// Mitsubishi GX Works2 project: ZhaoQing_FenRong_Debug   PLC: Q06UDEH (continued)

H750ImportCylinder2(ShuttleCarInOut:= H750ImportCylinder2IO );
ShuttleCarCurrentPosition( XCE OR XCD ,XCE ,XCD, FALSE, H750ImportCylinder2IO.iCurrentPos );
H750ImportCylinder2IO.xReady:=1;
H750ImportCylinder2IO.xForward:=M127;
H750ImportCylinder2IO.xBackward:=M128;
H750ImportCylinder2IO.xPosLimit:=1;
H750ImportCylinder2IO.xNegLimit:=1;
Y2BE:=H750ImportCylinder2IO.xCW;
Y2BD:=H750ImportCylinder2IO.xCCW;
H750ImportCylinder2IO.xCylinder:=1;

H750Conveyor5(ConveyorMotor:=H750Conveyor5IO);
H750Conveyor5IO.xForward:=M112;
H750Conveyor5IO.xCWPresent:=XB6;
Y2AC:=H750Conveyor5IO.xMotorCW;
H750Conveyor5IO.iDeviceID:=12131;

H750Conveyor6(ConveyorMotor:=H750Conveyor6IO);
H750Conveyor6IO.xForward:=M113;
H750Conveyor6IO.xCWPresent:=XB7;
Y2AD:=H750Conveyor6IO.xMotorCW;
H750Conveyor6IO.iDeviceID:=12132;
(********3巷道*************)
H750Switch3(ConveyorEntryIO:=H750Switch3ConveyorIn,
                         ConveyorExitIO:=H750Switch3ConveyorOut,
                        SwitchIO:=H750Switch3IO );
H750Switch3IO.xLiftCylinderExtendButton:=M129;
H750Switch3IO.xLiftCylinderRetractButton:=M130;
H750Switch3IO.xExitBarCylinderRetractButton:=M138;
Y2AF:=NOT (H750Switch3IO.xExitBarCylinderRetract OR m_iH750Switch3Select=2 );
Y2B1:=H750Switch3IO.xLiftCylinderExtend;
Y2B0:=H750Switch3IO.xLiftCylinderRetract;
H750Switch3IO.xLiftCylinderExtendDetect:=XBE;
H750Switch3IO.xLiftCylinderRetractDetect:=XBF;
H750Switch3ConveyorIn.xForward:=M131;
H750Switch3ConveyorIn.xCWPresent:=((m_iH750Switch3Select=1 OR m_iH750Switch3Select=0)  AND  XB9) OR (m_iH750Switch3Select=2 AND XC2);
Y2AB:=H750Switch3ConveyorIn.xMotorCW;
H750Switch3ConveyorIn.tLoadDelay:=T#3s;
H750Switch3ConveyorIn.iDeviceID:=12133;
H750Switch3ConveyorOut.xForward:=M132;
H750Switch3ConveyorOut.xCWPresent:=((m_iH750Switch3Select=1 OR m_iH750Switch3Select=0)  AND  XB9) OR (m_iH750Switch3Select=2 AND XC2);
Y2C0:=H750Switch3ConveyorOut.xMotorCW;
H750Switch3IO.xLiftCylinderExtendInit:=0;
H750Switch3ConveyorOut.iDeviceID:=12134;

H750ImportConveyor5(ConveyorMotor:=H750ImportConveyor5IO);
H750ImportConveyor5IO.xForward:=M133;
H750ImportConveyor5IO.xCWPresent:=XD1;
Y2BF:=H750ImportConveyor5IO.xMotorCW;
H750ImportConveyor5IO.tLoadDelay:=t#2S;
H750ImportConveyor5IO.iDeviceID:=12135;

H750ImportConveyor6(ConveyorMotor:=H750ImportConveyor6IO);
H750ImportConveyor6IO.xForward:=M134;
H750ImportConveyor6IO.xCWPresent:=XD3;
Y2C1:=H750ImportConveyor6IO.xMotorCW;
H750ImportConveyor6IO.tLoadDelay:=t#2S;
H750ImportConveyor6IO.iDeviceID:=12136;

H750ImportCylinder3(ShuttleCarInOut:= H750ImportCylinder3IO );
ShuttleCarCurrentPosition( XD4 OR XD5 ,XD5 ,XD4, FALSE, H750ImportCylinder3IO.iCurrentPos );
H750ImportCylinder3IO.xReady:=1;
H750ImportCylinder3IO.xForward:=M119;
H750ImportCylinder3IO.xBackward:=M120;
H750ImportCylinder3IO.xPosLimit:=1;
H750ImportCylinder3IO.xNegLimit:=1;
Y2C3:=H750ImportCylinder3IO.xCW;
Y2C2:=H750ImportCylinder3IO.xCCW;
H750ImportCylinder3IO.xCylinder:=1;
 (*******************************)
 (*<<<<<<<<<空框回流>>>>>>>>>>>>*)
 (*<<<<<<<<<1巷道>>>>>>>>>>>>*)
 H2500Export1Cylinder(ShuttleCarInOut:= H2500Export1CylinderIO );
ShuttleCarCurrentPosition( XDC OR XDD ,XDC ,XDD, FALSE, H2500Export1CylinderIO.iCurrentPos );
H2500Export1CylinderIO.xForward:=M147;
H2500Export1CylinderIO.xBackward:=M148;
Y2C8:=H2500Export1CylinderIO.xCW;
Y2C9:=H2500Export1CylinderIO.xCCW;
H2500Export1CylinderIO.xCylinder:=1;
H2500Export1CylinderIO.xPresentDetect1:=XDE;
H2500Export1CylinderIO.xPresentDetect2:=XDF;

H2500Export1Conveyor1(ConveyorMotor:=H2500Export1Conveyor1IO);
H2500Export1Conveyor1IO.xForward:=M149;
H2500Export1Conveyor1IO.xCWPresent:=XD8;
Y2C4:=H2500Export1Conveyor1IO.xMotorCW; 
H2500Export1Conveyor1IO.iDeviceID:=12137;
  
 H2500Export1Conveyor2(ConveyorMotor:=H2500Export1Conveyor2IO);
H2500Export1Conveyor2IO.xForward:=M150;
H2500Export1Conveyor2IO.xCWPresent:=XD9;
Y2C5:=H2500Export1Conveyor2IO.xMotorCW;
H2500Export1Conveyor2IO.iDeviceID:=12138;

 H2500Export1Conveyor3(ConveyorMotor:=H2500Export1Conveyor3IO);
H2500Export1Conveyor3IO.xForward:=M151;
H2500Export1Conveyor3IO.xCWPresent:=XDA;
Y2C6:=H2500Export1Conveyor3IO.xMotorCW;

 H2500Export1Conveyor4(ConveyorMotor:=H2500Export1Conveyor4IO);
H2500Export1Conveyor4IO.xForward:=M152;
H2500Export1Conveyor4IO.xCWPresent:=XDB;
Y2C7:=H2500Export1Conveyor4IO.xMotorCW;

 H2500Export1Switch(ConveyorEntryIO:= H2500Export1SwitchConveyorIn,
                         ConveyorExitIO:= H2500Export1SwitchConveyorOut,
                        SwitchIO:= H2500Export1SwitchIO );
H2500Export1SwitchIO.xLiftCylinderExtendButton:=M153;
H2500Export1SwitchIO.xLiftCylinderRetractButton:=M154;
Y2C8:=H2500Export1SwitchIO.xLiftCylinderExtend;
Y2C9:=H2500Export1SwitchIO.xLiftCylinderRetract;
H2500Export1SwitchIO.xLiftCylinderExtendDetect:=XBE;
H2500Export1SwitchIO.xLiftCylinderRetractDetect:=XBF;
H2500Export1SwitchConveyorIn.xForward:=M155;
H2500Export1SwitchConveyorIn.xCWPresent:=XDA OR XDB;
Y2D2:=H2500Export1SwitchConveyorIn.xMotorCW;
H2500Export1SwitchConveyorOut.xForward:=M156;
H2500Export1SwitchConveyorOut.xCWPresent:=XDA OR XDB;
(*Y2CD:=H2500Export1SwitchConveyorOut.xMotorCW;*)(*倍速链线体*)
H2500Export1SwitchIO.xLiftCylinderExtendInit:=1;

 (*<<<<<<<<<2巷道>>>>>>>>>>>>*)
  H2500Export2Cylinder(ShuttleCarInOut:= H2500Export2CylinderIO );
ShuttleCarCurrentPosition( XE4 OR XE5,XE4 ,XE5, FALSE, H2500Export2CylinderIO.iCurrentPos );
H2500Export2CylinderIO.xForward:=M157;
H2500Export2CylinderIO.xBackward:=M158;
Y2E0 :=H2500Export2CylinderIO.xCW;
Y2E1 :=H2500Export2CylinderIO.xCCW;
H2500Export2CylinderIO.xCylinder:=1;
H2500Export2CylinderIO.xPresentDetect1:=XE6;
H2500Export2CylinderIO.xPresentDetect2:=XE7;

H2500Export2Conveyor1(ConveyorMotor:=H2500Export2Conveyor1IO);
H2500Export2Conveyor1IO.xForward:=M159;
H2500Export2Conveyor1IO.xCWPresent:=XE0;
Y2CA:=H2500Export2Conveyor1IO.xMotorCW; 
  
 H2500Export2Conveyor2(ConveyorMotor:=H2500Export2Conveyor2IO);
H2500Export2Conveyor2IO.xForward:=M160;
H2500Export2Conveyor2IO.xCWPresent:=XE1;
Y2CB:=H2500Export2Conveyor2IO.xMotorCW;

 H2500Export2Conveyor3(ConveyorMotor:=H2500Export2Conveyor3IO);
H2500Export2Conveyor3IO.xForward:=M161;
H2500Export2Conveyor3IO.xCWPresent:=XE2;
Y2CC:=H2500Export2Conveyor3IO.xMotorCW;

 H2500Export2Conveyor4(ConveyorMotor:=H2500Export2Conveyor4IO);
H2500Export2Conveyor4IO.xForward:=M162;
H2500Export2Conveyor4IO.xCWPresent:=XE3;
Y2CD:=H2500Export2Conveyor4IO.xMotorCW;

 H2500Export2Switch(ConveyorEntryIO:= H2500Export2SwitchConveyorIn,
                         ConveyorExitIO:= H2500Export2SwitchConveyorOut,
                        SwitchIO:= H2500Export2SwitchIO );
H2500Export2SwitchIO.xLiftCylinderExtendButton:=M163;
H2500Export2SwitchIO.xLiftCylinderRetractButton:=M164;
Y2E0:=H2500Export2SwitchIO.xLiftCylinderExtend;
Y2E1:=H2500Export2SwitchIO.xLiftCylinderRetract;
H2500Export2SwitchIO.xLiftCylinderExtendDetect:=X102;
H2500Export2SwitchIO.xLiftCylinderRetractDetect:=X103;
H2500Export2SwitchConveyorIn.xForward:=M165;
H2500Export2SwitchConveyorIn.xCWPresent:=XE2 OR XE3;
Y2CC:=H2500Export2SwitchConveyorIn.xMotorCW;
H2500Export2SwitchConveyorOut.xForward:=M166;
H2500Export2SwitchConveyorOut.xCWPresent:=XE2 OR XE3;
(*Y2CD:=H2500Export1SwitchConveyorOut.xMotorCW;*)(*倍速链线体*)
H2500Export2SwitchIO.xLiftCylinderExtendInit:=1;
 (*<<<<<<<<<3巷道>>>>>>>>>>>>*)
 H2500Export3Cylinder(ShuttleCarInOut:= H2500Export3CylinderIO );
ShuttleCarCurrentPosition( XEC OR XED ,XEC ,XED, FALSE, H2500Export3CylinderIO.iCurrentPos );
H2500Export3CylinderIO.xForward:=M167;
H2500Export3CylinderIO.xBackward:=M168;
Y2D4:=H2500Export3CylinderIO.xCW;
Y2D5:=H2500Export3CylinderIO.xCCW;
H2500Export3CylinderIO.xCylinder:=1;
H2500Export3CylinderIO.xPresentDetect1:=XEE;
H2500Export3CylinderIO.xPresentDetect2:=XEF;

H2500Export3Conveyor1(ConveyorMotor:=H2500Export1Conveyor1IO);
H2500Export3Conveyor1IO.xForward:=M169;
H2500Export3Conveyor1IO.xCWPresent:=XE8;
Y2D0:=H2500Export3Conveyor1IO.xMotorCW; 
  
 H2500Export3Conveyor2(ConveyorMotor:=H2500Export1Conveyor2IO);
H2500Export3Conveyor2IO.xForward:=M170;
H2500Export3Conveyor2IO.xCWPresent:=XE9;
Y2D1:=H2500Export3Conveyor2IO.xMotorCW;

 H2500Export3Conveyor3(ConveyorMotor:=H2500Export1Conveyor3IO);
H2500Export3Conveyor3IO.xForward:=M171;
H2500Export3Conveyor3IO.xCWPresent:=XE9;
Y2D1:=H2500Export3Conveyor3IO.xMotorCW;

 H2500Export3Conveyor4(ConveyorMotor:=H2500Export1Conveyor4IO);
H2500Export3Conveyor4IO.xForward:=M172;
H2500Export3Conveyor4IO.xCWPresent:=XE9;
Y2D1:=H2500Export3Conveyor4IO.xMotorCW;

 H2500Export3Switch(ConveyorEntryIO:= H2500Export3SwitchConveyorIn,
                         ConveyorExitIO:= H2500Export3SwitchConveyorOut,
                        SwitchIO:= H2500Export3SwitchIO );
H2500Export3SwitchIO.xLiftCylinderExtendButton:=M173;
H2500Export3SwitchIO.xLiftCylinderRetractButton:=M174;
Y2D4:=H2500Export3SwitchIO.xLiftCylinderExtend;
Y2D5:=H2500Export3SwitchIO.xLiftCylinderRetract;
H2500Export3SwitchIO.xLiftCylinderExtendDetect:=XBE;
H2500Export3SwitchIO.xLiftCylinderRetractDetect:=XBF;
H2500Export3SwitchConveyorIn.xForward:=M175;
H2500Export3SwitchConveyorIn.xCWPresent:=XDA;
Y2D2:=H2500Export3SwitchConveyorIn.xMotorCW;
H2500Export3SwitchConveyorOut.xForward:=M176;
H2500Export3SwitchConveyorOut.xCWPresent:=XDA;
(*Y2CD:=H2500Export1SwitchConveyorOut.xMotorCW;*)(*倍速链线体*)
H2500Export3SwitchIO.xLiftCylinderExtendInit:=1;

(*倍速链二封车间顶升移载*)
H2500EmptyASwitch(ConveyorEntryIO:=H2500EmptyASwitchConveyorIn,
                                       ConveyorExitIO:=H2500EmptyASwitchConveyorOut,
                                       SwitchIO:=H2500EmptyASwitchIO);
H2500EmptyASwitchIO.xLiftCylinderExtendButton:=M97;
H2500EmptyASwitchIO.xLiftCylinderRetractButton:=M98;
Y256:=H2500EmptyASwitchIO.xLiftCylinderExtend;
Y255:=H2500EmptyASwitchIO.xLiftCylinderRetract;
H2500EmptyASwitchIO.xEntryBarCylinderRetractButton:=M106;
Y24F :=H2500EmptyASwitchIO.xEntryBarCylinderRetract;
H2500EmptyASwitchIO.xLiftCylinderExtendDetect:=X55;
H2500EmptyASwitchIO.xLiftCylinderRetractDetect:=X56;
H2500EmptyASwitchConveyorIn.xForward:=M99;
H2500EmptyASwitchConveyorIn.xCWPresent:=X4F;
(*Y248:=H2500EmptyASwitchConveyorIn.xMotorCW;*)
H2500EmptyASwitchConveyorOut.xForward:=M100;
H2500EmptyASwitchConveyorOut.xCWPresent:=X57;
Y257:=H2500EmptyASwitchConveyorOut.xMotorCW;

H2500EmptyBSwitch(ConveyorEntryIO:=H2500EmptyBSwitchConveyorIn,
                                       ConveyorExitIO:=H2500EmptyBSwitchConveyorOut,
                                       SwitchIO:=H2500EmptyBSwitchIO);
H2500EmptyBSwitchIO.xLiftCylinderExtendButton:=M101;
H2500EmptyBSwitchIO.xLiftCylinderRetractButton:=M102;
Y259:=H2500EmptyBSwitchIO.xLiftCylinderExtend;
Y258:=H2500EmptyBSwitchIO.xLiftCylinderRetract;
H2500EmptyBSwitchIO.xEntryBarCylinderRetractButton:=M107;
Y251:=H2500EmptyBSwitchIO.xEntryBarCylinderRetract;
H2500EmptyBSwitchIO.xLiftCylinderExtendDetect:=X58;
H2500EmptyBSwitchIO.xLiftCylinderRetractDetect:=X59;
H2500EmptyBSwitchConveyorIn.xForward:=M103;
H2500EmptyBSwitchConveyorIn.xCWPresent:=X52;
Y24A:=H2500EmptyBSwitchConveyorIn.xMotorCW;
H2500EmptyBSwitchConveyorOut.xForward:=M104;
H2500EmptyBSwitchConveyorOut.xCWPresent:=X5A;
Y25A:=H2500EmptyBSwitchConveyorOut.xMotorCW;
(*手动*)	
IF g_xManual OR g_xCommissioning THEN
	D3315:=0;
	D3140:=0;
	D3145:=0;
	D3320:=0;
	D3150 :=0;
	D3151 :=0;
	D3170:=0;
	D3171:=0;
	D3172:=0;
	D3190 :=0;
	D3191 :=0;
	D3192:=0;

END_IF;
(*自动*)	
IF g_xAuto AND NOT g_xCommissioning THEN
	(**************************上位机通讯数据************************)
	(*"分容入库前分流点
4004"	2315	5	分流方向	2315	"0：复位
1：读码失败
2：左排
3：右排"	3315	5	有板状态		1：无板，2：有板
*)
	IF NOT H2500BarCylinderIO.xEmpty THEN
		D3315:=2;
	ELSE
		D3315:=1;
	END_IF;
	H2500BarCylinderIO.iProductCategory:=D2315;
	(*"B1库入口
2009
（出入口编号1）"	2140	5	收到入库请求	2140	"1:复位
2:收到入库请求（只有在生成任务请求以后才置位）"	3140	5	入口状态	3140	"1：复位
2：入库请求"
*)
IF 	( (H2500RotorConveyorIO.xEmpty=0 AND H2500RotorConveyorIO.iProductCategory=3 AND H2500RotorIO.iCurrentPos=2) 
	OR (H2500RotorConveyorIO.xEmpty=0 AND H2500RotorConveyorIO.iProductCategory=2 AND H2500RotorIO.iCurrentPos=1))
	AND NOT M183
	THEN
	D3140:=2;
ELSE
	D3140:=1;
END_IF;
  H2500RotorConveyorIO.xPutInto:=M69;(*转台取料后复位*)(*触摸屏上制作强制完成按钮*)
 m_tpH2500RotorReset(IN:= D2141 = 2 AND NOT H2500RotorConveyorIO.xCCWPresent AND NOT H2500RotorConveyorIO.xCWPresent AND NOT X134 ,
 											PT:= t#3S ,
 											Q:= M69 ,
 											ET:= m_tH2500RotorResetCurrentTime);
(*IF LDP(TRUE, D2141 = 2 AND NOT H2500RotorConveyorIO.xCCWPresent AND NOT H2500RotorConveyorIO.xCWPresent AND NOT X134) THEN
	M69:=1;
ELSE
	M69:=0;
END_IF;*)
(*取货完成，m69，H2500RotorConveyorIO.xPutInto*)
(*"B1库出口
2010
（出入口编号1）"	2145	5	出库完成状态	2145	"1：复位
2：出库完成 "	3145	5	出口状态	3145	"1:复位
2:允许出库"
*)
IF H750RotorIO.iCurrentPos=2
	AND H750RotorConveyorIO.xEmpty  
	AND NOT H750RotorConveyorIO.xCCWPresent 
	AND NOT H750RotorConveyorIO.xCWPresent
	AND NOT M179   THEN
	D3145:=2;
ELSE
	D3145:=1;
END_IF;
H750RotorConveyorIO.xPutInto:=M144;(*触摸屏上制作强制完成按钮人工在转台上上料入常温库*)
IF D2145=2 THEN
	M144:=1;
ELSE
	M144:=0;
END_IF;
(*出库转台旋转方向*)
IF D2146=2 THEN
	m_xH750RotorDirection:=1;
ELSE
	m_xH750RotorDirection:=0;
END_IF;

(*"常温入库前分流（分容后）
4005"	2320	5	分流方向	2320	"0：复位
1：读码失败
2：流向C1库，
3：流向C2库
4：流向C3库
5:等待"	3320	5	有板状态	3320	1：无板，2：有板
*)
IF H750Conveyor1IO.xEmpty=0 THEN
	D3320:=2;
ELSE
	D3320:=1;
END_IF;

H750Conveyor1IO.iProductCategory:=D2320;

(*"C1库入口(分容后）
2011
（出入口编号1）"	2150	5				3150	5	位置1有板状态	3150	1：无板，2：有板
								位置2有板状态	3151	1：无板，2：有板
								手动入库请求	3152	1:复位，2：请求入库
*)
IF H750ImportCylinder1IO.iCurrentPos=2 AND XC8 AND NOT M180  THEN
	D3150 :=2;
ELSIF M180 THEN (*禁止入库*)
	D3150 :=0;
ELSE
	D3150 :=1;	
END_IF;
IF H750ImportCylinder1IO.iCurrentPos=2  AND XC9 AND NOT M180 THEN
	D3151 :=2;
ELSIF M180 THEN(*禁止入库*)
	D3151 :=0;
ELSE
	D3151 :=1;	
END_IF;
IF g_xImport1Force THEN
	D3152:=2;
ELSE
	D3152:=1;
END_IF;
(*3170	5	位置1有板状态	3170	1：无板，2：有板
		位置2有板状态	3171	1：无板，2：有板
		手动入库请求	3172	1:复位，2：请求入库*)
IF H750ImportCylinder2IO.iCurrentPos=2 AND XCF AND NOT M181  THEN
	D3170 :=2;
ELSIF  M181 THEN(*禁止入库*)
	D3170 :=0;
ELSE
	D3170 :=1;	
END_IF;
IF H750ImportCylinder2IO.iCurrentPos=2  AND XD0 AND NOT M181 THEN
	D3171 :=2;
ELSIF M181 THEN(*禁止入库*)
	D3171 :=0;
ELSE
	D3171 :=1;	
END_IF;
IF g_xImport2Force THEN
	D3172:=2;
ELSE
	D3172:=1;
END_IF;		
(*"C3库入口(分容后）
2019
（出入口编号1）"	2190	5				3190	5	位置1有板状态	3190	1：无板，2：有板
								位置2有板状态	3191	1：无板，2：有板
								手动入库请求	3192	1:复位，2：请求入库
*)
IF H750ImportCylinder3IO.iCurrentPos=2 AND XD6 AND NOT M182  THEN
	D3190 :=2;
ELSIF M182 THEN(*禁止入库*)
	D3190 :=0;
ELSE
	D3190 :=1;	
END_IF;
IF H750ImportCylinder3IO.iCurrentPos=2  AND XD7 AND NOT M182 THEN
	D3191 :=2;
ELSIF M182 THEN(*禁止入库*)
	D3191 :=0;
ELSE
	D3191 :=1;	
END_IF;
IF g_xImport3Force THEN
	D3192:=2;
ELSE
	D3192:=1;
END_IF;	

	(*****************************二封车间RGV控制******************************)
	
	(*****************************二封4号机机对接信号******************************)	
	QuarPackage4Stub.xUnloadRequestAkn:=X120;
	QuarPackage4Stub.xLoadRequest:=X122;	
	Y2FA:=QuarPackage4Stub.xUnloadRequest;(*X10CD*)
	Y2F8:=QuarPackage4Stub.xLoadRequestAkn;(*X10CE*)
	
	H850Conveyor2IOTrans.xLoad:=QuarPackage4Stub.xLoadRequest;
	QuarPackage4Stub.xLoadRequestAkn:=H850Conveyor2IOTrans.xEmpty;
	H850Conveyor1IOTrans.xUnload:=QuarPackage4Stub.xUnloadRequestAkn;
	QuarPackage4Stub.xUnloadRequest:=NOT H850Conveyor1IOTrans.xEmpty;
	
	H850Conveyor2IOTrans.xPutInto:=NOT H850Conveyor2IOTrans.xBusy AND SM412;
	H850Conveyor1IOTrans.xPutInto:=NOT H850Conveyor1IOTrans.xBusy AND SM412;
	(*****************************二封3号机机对接信号******************************)	
	QuarPackage3Stub.xUnloadRequestAkn:=X124;
	QuarPackage3Stub.xLoadRequest:=X126;	
	Y2FE:=QuarPackage3Stub.xUnloadRequest;(*X10CD*)
	Y2FC:=QuarPackage3Stub.xLoadRequestAkn;(*X10CE*)

	H850Conveyor4IOTrans.xLoad:=QuarPackage3Stub.xLoadRequest;
	QuarPackage3Stub.xLoadRequestAkn:=H850Conveyor4IOTrans.xEmpty;
	H850Conveyor3IOTrans.xUnload:=QuarPackage3Stub.xUnloadRequestAkn;
	QuarPackage3Stub.xUnloadRequest:=NOT H850Conveyor3IOTrans.xEmpty;

	H850Conveyor4IOTrans.xPutInto:=NOT H850Conveyor4IOTrans.xBusy AND SM412;
	H850Conveyor3IOTrans.xPutInto:=NOT H850Conveyor3IOTrans.xBusy AND SM412;
	(*****************************二封2号机机对接信号******************************)	
	QuarPackage2Stub.xUnloadRequestAkn:=X128;
	QuarPackage2Stub.xLoadRequest:=X12A;	
	Y302:=QuarPackage2Stub.xUnloadRequest;(*X10CD*)
	Y300:=QuarPackage2Stub.xLoadRequestAkn;(*X10CE*)
	
	H850Conveyor6IOTrans.xLoad:=QuarPackage2Stub.xLoadRequest;
	QuarPackage2Stub.xLoadRequestAkn:=H850Conveyor6IOTrans.xEmpty;
	H850Conveyor5IOTrans.xUnload:=QuarPackage2Stub.xUnloadRequestAkn;
	QuarPackage2Stub.xUnloadRequest:=NOT H850Conveyor5IOTrans.xEmpty;
	(*自动复位程序*)
	H850Conveyor6IOTrans.xPutInto:=NOT H850Conveyor6IOTrans.xBusy AND SM412;
	H850Conveyor5IOTrans.xPutInto:=NOT H850Conveyor5IOTrans.xBusy AND SM412;
	(*****************************二封1号机机对接信号******************************)	
		QuarPackage1Stub.xUnloadRequestAkn:=X12C;
	QuarPackage1Stub.xLoadRequest:=X12E;	
	Y306:=QuarPackage1Stub.xUnloadRequest;(*X10CD*)
	Y304:=QuarPackage1Stub.xLoadRequestAkn;(*X10CE*)

	H850Conveyor8IOTrans.xLoad:=QuarPackage1Stub.xLoadRequest;
	QuarPackage1Stub.xLoadRequestAkn:=H850Conveyor8IOTrans.xEmpty;
	H850Conveyor7IOTrans.xUnload:=QuarPackage1Stub.xUnloadRequestAkn;
	QuarPackage1Stub.xUnloadRequest:=NOT H850Conveyor7IOTrans.xEmpty;
		(*自动复位程序*)
	H850Conveyor8IOTrans.xPutInto:=NOT H850Conveyor8IOTrans.xBusy AND SM412;
	H850Conveyor7IOTrans.xPutInto:=NOT H850Conveyor7IOTrans.xBusy AND SM412;
	(*****************************二封与RGV对接信号******************************)
	(*发送*)
   D221:=QuarPackageRGV.iDestinationPos;	
   D222.0:=QuarPackageRGV.xAuto; 	
   D222.1:=QuarPackageRGV.xMdiExe;
   D222.2:=QuarPackageRGV.xLoad1;
   D222.3:=QuarPackageRGV.xUnload1;
   D222.4:=H850Conveyor1IOTrans.xEmpty;
   D222.5:=H850Conveyor2IOTrans.xEmpty;
   D222.6:=H850Conveyor3IOTrans.xEmpty;
   D222.7:=H850Conveyor4IOTrans.xEmpty;
   D222.8:=H850Conveyor5IOTrans.xEmpty;
   D222.9:=H850Conveyor6IOTrans.xEmpty;
   D222.A:=H850Conveyor7IOTrans.xEmpty;
   D222.B:=H850Conveyor8IOTrans.xEmpty;
   D222.C:=H850Switch2ConveyorIn.xEmpty;
   D222.D:=H850Switch3ConveyorIn.xEmpty;
   
   D223.0:=QuarPackageRGV.xRemoteReset;
   D223.1:=H850Conveyor1IOTrans.xNextRun;
   D223.2:=H850Conveyor2IOTrans.xNextRun;
   D223.3:=H850Conveyor3IOTrans.xNextRun;
   D223.4:=H850Conveyor4IOTrans.xNextRun;  
   D223.5:=H850Conveyor5IOTrans.xNextRun;
   D223.6:=H850Conveyor6IOTrans.xNextRun;
   D223.7:=H850Conveyor7IOTrans.xNextRun;
   D223.8:=H850Conveyor8IOTrans.xNextRun;  
   D223.9:=H850Switch3ConveyorOut.xNextRun; 
   QuarPackageRGV.xRemoteReset:=M191;
   QuarPackageRGV.xAuto:=M186;
   (*接收*)
   QuarPackageRGV.iCurrentPostion:=D421;
   QuarPackageRGV.xMdiDone:=D422.0;
   QuarPackageRGV.xEmpty1:=D422.1;
   QuarPackageRGV.xNextRun1:=D422.2;
   QuarPackageRGV.xEmpty2:=D422.3;
   QuarPackageRGV.xNextRun2:=D422.4;
   H850Conveyor1IOTrans.xLoad:= D422.5;
   H850Conveyor3IOTrans.xLoad:= D422.6; 
   H850Conveyor5IOTrans.xLoad:= D422.7; 
   H850Conveyor7IOTrans.xLoad:= D422.8;
    H850Conveyor2IOTrans.xUnload:= D422.9;
   H850Conveyor4IOTrans.xUnload:= D422.A; 
   H850Conveyor6IOTrans.xUnload:= D422.B; 
   H850Conveyor8IOTrans.xUnload:= D422.C;  
  (** H850Switch2IO.xEntryEnable:=D422.D*)
   H850Switch2IO.xEntryEnable:=D422.D;
   H850Switch3IO.xExitEnable:=D422.E;
   QuarPackageRGV.xCollisionAlarm:=D423.0;
	
   
      (*去分容库位置*)
    IF M185 THEN
   	QuarPackageRGV.xMdiExe:=1;
   	QuarPackageRGV.iDestinationPos:=5;
    END_IF;   
       (*1号上料*)
   IF M187 THEN
   	QuarPackageRGV.xMdiExe:=1;
   	QuarPackageRGV.iDestinationPos:=4;
   END_IF;
       (*2号上料*)
     IF M188 THEN
   	QuarPackageRGV.xMdiExe:=1;
   	QuarPackageRGV.iDestinationPos:=3;
     END_IF; 
         (*3号上料*)
    IF M189 THEN
   		QuarPackageRGV.xMdiExe:=1;
   		QuarPackageRGV.iDestinationPos:=2;
    END_IF;
          (*4号上料*)
   IF M190 THEN
   	QuarPackageRGV.xMdiExe:=1;
   	QuarPackageRGV.iDestinationPos:=1;
   END_IF;   	
   	
	(*=============================================*)
	(*****************************上料去分容库******************************)	
	H850Switch2IO.xLiftCylinderExtendInit:=0;
(*	IF  M880 OR X69  THEN
		H850Switch2IO.xEntryEnable:=1;
	ELSE
		H850Switch2IO.xEntryEnable:=0;
	END_IF;*)
	IF M880 OR X69 THEN
		m_xManualLoad:=1;(*人工上料任务*)
	END_IF;
	H850Switch4Task(xCondition1:=NOT  H850Conveyor14IO.xEmpty ,
									xCondition2:=m_xManualLoad,
									xCondition3:=FALSE ,
									xCondition4:=FALSE ,
									xCondition5:= FALSE ,
									xTaskComplete:= LDP(TRUE,H850Switch4ConveyorOut.xEmpty) ,
									xReset:= g_xResetSingle AND g_iDeviceIDSelect=12301 ,
									iPriority:= m_iH850Switch4Task );
	IF m_iH850Switch4Task=2 THEN
		H850Conveyor12IO.xLoad:=1;
	END_IF;
	IF H850Conveyor12IO.xBusy THEN
		H850Conveyor12IO.xLoad:=0;
	END_IF;
	IF LDF(TRUE,H850Conveyor12IO.xEmpty) THEN
		m_xManualLoad:=0;
	END_IF;
	H850CONVEYOR12IO.tLoadDelay:=T#1s500ms;
	H850Switch4IO.xSwithEnable:=1;
	H850Switch4IO.xLiftCylinderExtendInit:=m_iH850Switch4Task<>1;
	H850Switch4ConveyorOut.xUnload:=H850CONVEYOR1iO.xEmpty;
	IF X136 OR g_xPassQualityDetectStation1  THEN(*品检按钮盒*)
		m_xDefectDetect1Complete:=1;
	END_IF;
	IF LDF(TRUE,H850conveyor13IO.xEmpty) THEN
		m_xDefectDetect1Complete:=0;
	END_IF;
	h850Switch2IO.xSwithEnable:=1;
	(*品检工位1*)
	H850Switch2IO.xExitEnable:=H850conveyor13IO.xEmpty AND m_xDefectDetect1Complete;
	H850Conveyor13IO.xLoad:=H850Switch2ConveyorOut.xNextRun;
	(*品检工位2*)	
	IF X137 OR g_xPassQualityDetectStation2 THEN
		m_xDefectDetect2Complete:=1;
	END_IF;
	IF LDF(TRUE,H850Switch5ConveyorIn.xEmpty) THEN
		m_xDefectDetect2Complete:=0;
	END_IF;	
	H850Conveyor13IO.xUnload:=H850Switch5ConveyorIn.xEmpty AND H850Conveyor14IO.xEmpty AND m_xDefectDetect2Complete ;
	H850Switch5IO.xEntryEnable:=H850Conveyor13IO.xNextRun;
	H850Switch5IO.xLiftCylinderExtendInit:=h850Conveyor14IO.xEmpty;
	H850Switch5IO.xSwithEnable:=1;
	H850Switch5ConveyorIn.tLoadDelay:=T#1s500ms;
	H850Switch5IO.xExitEnable:=H850CONVEYOR14iO.xEmpty;
	(*品检工位3*)	
	IF X13A OR g_xPassQualityDetectStation3 THEN
		m_xDefectDetect3Complete:=1;
	END_IF;
	IF LDF(TRUE,H850Switch4ConveyorOut.xEmpty) THEN
		m_xDefectDetect3Complete:=0;
	END_IF;	
	h850Conveyor14IO.xLoad:=H850Switch5ConveyorOut.xNextRun ;
(*	H850Switch5IO.xExitEnable:=H850CONVEYOR1iO.xEmpty;*)
	H850Conveyor14IO.xUnload:=H850Switch4ConveyorOut.xEmpty AND m_iH850Switch4Task=1 AND m_xDefectDetect3Complete;
	H850Switch4ConveyorOut.xLoad:=H850Conveyor14IO.xNextRun;
	H850Conveyor1IO.xLoad:=H850Switch4ConveyorOut.xNextRun;
	
	IF ldp(TRUE,H850Switch2ConveyorOut.xEmpty) THEN   (*上料计数*)
		D20:=D20+1;
	END_IF;
	IF M88 THEN(*计数清零*)
		D20:=0;
	END_IF;
	
	
	IF COnveyor7IO.xEmpty THEN
		Lifter7IO.xMDIExe:=1;
		Lifter7Io.iDestinationPos:=1;
	END_IF;
	IF conveyor7IO.xEmpty=0 THEN
		Lifter7Io.xMDIExe:=1;
		Lifter7io.iDestinationPos:=2;
	END_IF;
	IF Lifter7IO.iCurrentPos=1 THEN
		H850Conveyor1IO.xUnload:=COnveyor7IO.xEmpty  
		                                                    AND NOT g_xForbidLifter7 (*提升机7禁止入料*)
		                                                    AND NOT Conveyor7IO.xOverWidthAlarm;(*提升机7超宽检测*)
	ELSE
		H850Conveyor1IO.xUnload:=0;
	END_IF;
		COnveyor7IO.xLoad:=H850Conveyor1IO.xNextRun;
		IF Lifter7IO.iCurrentPos=2 THEN
			COnveyor7IO.xUnload:=H2500Conveyor1IO.xEmpty;
		ELSE 
			COnveyor7IO.xUnload:=0;
		END_IF;
		H2500Conveyor1IO.xLoad:=COnveyor7IO.xNextRun;
		H2500SwitchIO.xLiftCylinderExtendInit:=1;
		h2500SwitchIO.xSwithEnable:=1;
		h2500Conveyor1IO.xUnload:=H2500SwitchConveyorIn.xEmpty AND H2500SwitchConveyorOut.xEmpty AND H2500BarCylinderIO.xEmpty;
		H2500SwitchIO.xEntryEnable:=H2500Conveyor1IO.xNextRun;
		H2500SwitchIO.xExitEnable:=H2500BarCylinderIO.xEmpty;
		Y282:=H2500BarCylinderIO.xEmpty;(*前挡停器，不为空的时候顶起*)
		IF H2500RotorIO.iCurrentPos=1 AND (H2500BarCylinderIO.iProductCategory=2 OR H2500BarCylinderIO.iProductCategory=3)  THEN			
			H2500BarCylinderIO.xUnload:=H2500RotorConveyorIO.xEmpty;
		ELSE
			H2500BarCylinderIO.xUnload:=0;
		END_IF;
	    H2500RotorConveyorIO.xLoad:=H2500BarCylinderIO.xNextRun;   
	    IF LDP(TRUE,H2500BarCylinderIO.xNextRun) THEN
	    	H2500RotorConveyorIO.iProductCategory:= H2500BarCylinderIO.iProductCategory;
	    	END_IF;
		IF H2500RotorConveyorIO.xEmpty=0 AND H2500RotorConveyorIO.iProductCategory=3 THEN
			H2500RotorIO.xMDIExe:=1;
			H2500RotorIO.iDestinationPos:=2;
		ELSE
			H2500RotorIO.xMDIExe:=1;
			H2500RotorIO.iDestinationPos:=1;			
		END_IF;	

         (*分容出库，常温库入库*)
       IF H750RotorConveyorIO.xEmpty THEN
       	H750RotorIO.xMDIExe:=1;
       	H750RotorIO.iDestinationPos:=2;
       END_IF;
         IF H750RotorConveyorIO.xEmpty=0 AND m_xH750RotorDirection THEN
       	H750RotorIO.xMDIExe:=1;
       	H750RotorIO.iDestinationPos:=1;
         ELSIF H750RotorConveyorIO.xEmpty=0 AND NOT m_xH750RotorDirection THEN
         H750RotorIO.xMDIExe:=1;
       	H750RotorIO.iDestinationPos:=3;       	
         END_IF;     
         IF  H750RotorIO.iCurrentPos=1 THEN
         	H750RotorConveyorIO.xUnload:=H750SwitchConveyorIn.xEmpty;
         	H750SwitchIO.xEntryEnable:=H750RotorConveyorIO.xNextRun;
         	H750RotorConveyorIO.xUnloadCCW:=1;
	     ELSIF H750RotorIO.iCurrentPos=3 THEN
          	H750RotorConveyorIO.xUnload:=H750SwitchConveyorIn.xEmpty;
         	H750SwitchIO.xEntryEnable:=H750RotorConveyorIO.xNextRun;
         	H750RotorConveyorIO.xUnloadCCW:=0;        	
         ELSE
         	H750RotorConveyorIO.xUnload:=0;
         	H750SwitchIO.xEntryEnable:=0;
         	H750SwitchConveyorIn.xLoad:=0;
         END_IF;
         H750SwitchIO.xSwithEnable:=1;
         H750SwitchIO.xExitEnable:=H750Conveyor1IO.xEmpty;
         H750Conveyor1IO.xLoad:=H750SwitchConveyorOut.xNextRun;
         (*条码扫描结果，显示分配的巷道，写在了传输线块的产品类型里面了，通过一段一段的传输线传输下去*)
         IF  H750Conveyor1IO.iProductCategory=2 OR H750Conveyor1IO.iProductCategory=3 OR H750Conveyor1IO.iProductCategory=4  THEN
         	H750Conveyor1IO.xUnload:=H750Conveyor2IO.xEmpty;
         ELSE
         	H750Conveyor1IO.xUnload:=0;
         END_IF;	
         	H750Conveyor2IO.xLoad:=H750Conveyor1IO.xNextRun;
         	(*分流信息传递*)
         	IF ldp(TRUE, H750Conveyor1IO.xNextRun) THEN
         		H750Conveyor2IO.iProductCategory:=H750Conveyor1IO.iProductCategory;
         	END_IF;
         	(*触摸屏上计数程序*)
         	IF LDP(TRUE,H750Conveyor2IO.xEmpty=0) THEN
         		D22:=D22+1;
         	END_IF;
         	IF M140 THEN
         		D22:=0;
         	END_IF;
         	(**********************************)
           H750Conveyor2IO.xUnload:=H750Switch1ConveyorIn.xEmpty AND H750Conveyor2IO.iProductCategory<>0 ;
           H750Switch1IO.xEntryEnable:=H750Conveyor2IO.xNextRun;
           (*分流信息传递到巷道1的顶升移载处*)
           IF LDP(TRUE,H750Conveyor2IO.xNextRun) THEN
           	H750Switch1ConveyorIn.iProductCategory:=H750Conveyor2IO.iProductCategory;
           END_IF;
           (*分流信息显示为本巷道，启动顶升移载*)
           IF H750Switch1ConveyorIn.iProductCategory=2 THEN
           	H750Switch1IO.xSwithEnable:=1;
           ELSE
           	H750Switch1IO.xSwithEnable:=0;
           END_IF;
           (*双料入库，优先选择1 ，当1结束后恢复到0，2秒 ，然后再跳到2,0状态用来复位移载的出料*) 
           m_tonSwitch1NOSeleteDelay(IN:= m_iH750Switch1Select=0 ,PT:= t#2S ,Q:=m_xSwitch1NoSeleteDelay,ET:= m_tSwitch1NOSeleteDelayCurrentTi );
         IF   m_xSwitch1NoSeleteDelay THEN
         	m_xSwitch1SeleteDelay:=1;
         END_IF;
         IF ldf(TRUE, H750ImportConveyor1IO.xEmpty)  OR ldf(TRUE,H750ImportConveyor2IO.xEmpty) THEN
         	m_xSwitch1SeleteDelay:=0;
         END_IF;
   (*        m_tonSwitch1SeleteDelay(IN:= m_xSwitch1NOSeleteDelay  ,PT:= t#10S ,Q:= m_xSwitch1SeleteDelay ,ET:= m_tSwitch1SeleteDelayCurrentTime );     *)      
           IF H750ImportConveyor1IO.xEmpty AND  m_xSwitch1SeleteDelay   THEN
           		m_iH750Switch1Select:=1;
	           	ELSIF NOT H750ImportConveyor1IO.xEmpty AND H750ImportConveyor2IO.xEmpty AND m_xSwitch1SeleteDelay  THEN
           	  	m_iH750Switch1Select:=2;
          	 ELSE
           		m_iH750Switch1Select:=0;
           END_IF;
           IF H750Switch1IO.xSwithEnable THEN
         	  H750Switch1io.xExitEnable:=((H750ImportConveyor1IO.xEmpty AND m_iH750Switch1Select=1) 
                                                          OR   (H750ImportConveyor2IO.xEmpty AND m_iH750Switch1Select=2)) AND H750ImportCylinder1IO.iCurrentPos=1;
           ELSE
   	        	H750Switch1io.xExitEnable:= H750Conveyor3IO.xEmpty AND H750Switch1ConveyorIn.iProductCategory>2;
    	        H750Conveyor3IO.xLoad:= H750Switch1ConveyorIn.xNextRun ;
            END_IF;
           	                                          
           H750ImportConveyor1IO.xLoad:=H750Switch1ConveyorOut.xNextRun AND m_iH750Switch1Select=1 ;
   	       H750ImportConveyor2IO.xLoad:=H750Switch1ConveyorOut.xNextRun AND m_iH750Switch1Select=2 ;
   	       IF  H750ImportConveyor1IO.xEmpty =0 AND H750ImportConveyor2IO.xEmpty =0 AND XC8 AND XC9 THEN
   	       	H750ImportCylinder1IO.xMDIExe:=1;
   	       	H750ImportCylinder1IO.iDestinationPos:=2;
   	       	H750ImportConveyor1IO.xPutInto:=0;
   	       	H750ImportConveyor2IO.xPutInto:=0;
   	       END_IF;
   	       IF g_xImport1Force THEN (* 1巷道单框强制入库*)
   	       	H750ImportCylinder1IO.xMDIExe:=1;
   	       	H750ImportCylinder1IO.iDestinationPos:=2;
   	       	H750ImportConveyor1IO.xPutInto:=0;
   	       	H750ImportConveyor2IO.xPutInto:=0;   
   	       	END_IF;	       	
   	       IF NOT XC8 AND NOT XC9 THEN
   	       		H750ImportCylinder1IO.xMDIExe:=1;
   	       		H750ImportCylinder1IO.iDestinationPos:=1;
   	       END_IF;
   	       IF LDP(TRUE,H750ImportCylinder1IO.iCurrentPos=1 AND NOT H750ImportConveyor1IO.xCWPresent AND NOT H750ImportConveyor2IO.xCWPresent) THEN   	       	
   	       		H750ImportConveyor1IO.xPutInto:=1;
   	       		H750ImportConveyor2IO.xPutInto:=1;
   	       END_IF;
  (***************2 巷道****************) 
  			IF LDP(TRUE,H750Switch1ConveyorIn.xNextRun) THEN
  				H750Conveyor3IO.iProductCategory:= H750Switch1ConveyorIn.iProductCategory;  
  			END_IF;
         	H750Conveyor3IO.xUnload:=H750Conveyor4IO.xEmpty AND H750Conveyor3IO.iProductCategory>2 ;
         	H750Conveyor4IO.xLoad:=H750Conveyor3IO.xNextRun;
         	H750Conveyor4IO.xUnload:=H750Switch2ConveyorIn.xEmpty AND H750Conveyor4IO.iProductCategory>2 ;
   			IF LDP(TRUE,H750Conveyor3IO.xNextRun) THEN
  				H750Conveyor4IO.iProductCategory:= H750Conveyor3IO.iProductCategory;  
  			END_IF;             
            H750Switch2IO.xEntryEnable:=H750Conveyor4IO.xNextRun;
           (*分流信息传递到巷道2的顶升移载处*)
           IF LDP(TRUE,H750Conveyor4IO.xNextRun) THEN
           	H750Switch2ConveyorIn.iProductCategory:=H750Conveyor4IO.iProductCategory;
           END_IF;
           (*分流信息显示为本巷道，启动顶升移载*)
           IF H750Switch2ConveyorIn.iProductCategory=3 THEN
           	H750Switch2IO.xSwithEnable:=1;
           ELSE
           	H750Switch2IO.xSwithEnable:=0;
           END_IF;
           (*双料入库，优先选择1 ，当1结束后恢复到0，2秒 ，然后再跳到2,0状态用来复位移载的出料*) 
          m_tonSwitch2NOSeleteDelay(IN:= m_iH750Switch2Select=0 ,PT:= t#2S ,Q:=m_xSwitch2NoSeleteDelay,ET:= m_tSwitch2NOSeleteDelayCurrentTi);
         IF   m_xSwitch2NoSeleteDelay THEN
         	m_xSwitch2SeleteDelay:=1;
         END_IF;
         IF ldf(TRUE, H750ImportConveyor3IO.xEmpty)  OR ldf(TRUE,H750ImportConveyor4IO.xEmpty) THEN
         	m_xSwitch2SeleteDelay:=0;
         END_IF;
   (*        m_tonSwitch1SeleteDelay(IN:= m_xSwitch1NOSeleteDelay  ,PT:= t#10S ,Q:= m_xSwitch1SeleteDelay ,ET:= m_tSwitch1SeleteDelayCurrentTime );     *)      
           IF H750ImportConveyor3IO.xEmpty AND  m_xSwitch2SeleteDelay   THEN
           		m_iH750Switch2Select:=1;
	           	ELSIF NOT H750ImportConveyor3IO.xEmpty AND H750ImportConveyor4IO.xEmpty AND m_xSwitch2SeleteDelay  THEN
           	  	m_iH750Switch2Select:=2;
          	 ELSE
           		m_iH750Switch2Select:=0;
           END_IF;
           IF H750Switch2IO.xSwithEnable THEN
         	  H750Switch2io.xExitEnable:=((H750ImportConveyor3IO.xEmpty AND m_iH750Switch2Select=1) 
                                                          OR   (H750ImportConveyor4IO.xEmpty AND m_iH750Switch2Select=2)) AND  H750ImportCylinder2IO.iCurrentPos=1;